VERSION : 1.0
// Support: tech.team.motioncontrol@siemens.com
   VAR_INPUT
      Cfg_EventListOffset : Int;   // Commanded event list offset (used for scrolling)
      Cfg_FilterCategory : Int;   // Filtered category number
      Cfg_TimeSortDirection : Bool;   // 1=newest first; 0=oldest first
      Cmd_FilterActiveEvents : Bool;   // 1=only show active events; 0=show all events
      Cmd_FilterCategory : Bool;   // Filter events to show only selected category number
      Cmd_SortCategory : Bool;   // 1=Sort events by ascending category number
   END_VAR
   VAR_OUTPUT
      Sts_EventListOffset : Int;   // Actual event list offset
      Sts_FilterExcludedNumEvents : Int;   // The number of events excluded by filtering
      Sts_SortFilterNumEvents : Int;   // Number of events in the sorted or filtered event list
   END_VAR
   VAR_IN_OUT
      In_Events : Array[0.."CPG_NO_OF_STS_ELEMENTS_EVENT_SUM_UPPER_LIM"] of "CPG_typeEvent";   // Input Event list to be sorted and/or filtered
      In_NumEvents : Int;   // Number of events to be sorted and/or filtered
      Sts_SortFilterEventList : Array[0.."CPG_NO_OF_HMI_SORT_EVENTS_UPPER_LIM"] of "CPG_typeEvent";   // Output sorted and/or filtered event list
   END_VAR
   VAR
      statFirstScan : Bool;   // stat first scan bit
      statCatIndex : Int;   // stat category index
      statCopiedIndex : Int;   // stat copied index
      statFilterActive : Bool;   // stat filter active = 1
      statFilterCategory : Bool;   // stat filter category
      statFilteredIndex : Int;   // stat filtered index
      statIndex : Int;   // stat index
      statLocalEventOffset : Int;   // stat local event offset
      statMaxInputSize : Int;   // stat max input size
      statMaxLocalInputSize : Int;   // stat max local input size
      statMaxOutputSize : Int;   // stat max output size
      statMaxParameterInputSize : Int;   // stat max parameter input size
      statNumDisplayedEvents : Int;   // stat num displayed events
      statNumFilteredEvents : Int;   // stat num of filtered events
      statPrevNumEvents : Int;   // stat previous number of events
      statSortedIndex : Int;   // stat sorted index
      statFilteredEventList : Array[0.."CPG_NO_OF_STS_ELEMENTS_EVENT_SUM_UPPER_LIM"] of "CPG_typeEvent";   // stat sorted event list
      statZeroEvent : "CPG_typeEvent";   // stat zeroized event list
   END_VAR
   VAR_TEMP
      tempMoveBlkVariantRetVal : Int;   // temp return value for BlockMoveVariant
   END_VAR
   VAR CONSTANT
      ZERO_VALUE : Int := 0;
   END_VAR
BEGIN
   //============================================================================================================
   // SIEMENS AG
   // (c)Copyright 2018 All Rights Reserved
   //------------------------------------------------------------------------------------------------------------
   // Project: CPG Template
   // Tested with: S7-1500 with FW version V2.1
   // Engineering: TIA Portal V14
   // Restrictions: ---
   // Requirements: S7-1500
   // Functionality: Control Event Sort Filter commands
   // Support: tech.team.motioncontrol@siemens.com
   //------------------------------------------------------------------------------------------------------------
   // Change log table:
   // Version       Date               Expert in charge    Changes applied
   //  01.00.00     01.01.2018         MP                  Initial Release & PackML V2.1  Renamed CPG V1.0
   //  01.01.00     29.05.2018         JP                  Adopted to styleguide
   //============================================================================================================
   // Function : CPG_EventSortFilter
   //============================================================================================================

   IF #statFirstScan = FALSE THEN
       // initialize & determine max array size
       // input array size (i.e. Array[0.."CPG_NO_STS_ELEMENTS_EVENT_STATUS"] of "typeCPG_Event")
       "CPG_ArrayLength"(arrayToBeSized := #In_Events,
                         arraySize => #statMaxParameterInputSize);

       //output array size for HMI (i.e. Array[0.."CPG_NO_HMI_SORT_EVENTS"] of "typeCPG_Event")
       "CPG_ArrayLength"(arrayToBeSized := #Sts_SortFilterEventList,
                         arraySize => #statMaxOutputSize);

       // internal/temporary array size (i.e. Array[0.."CPG_NO_STS_ELEMENTS_EVENT_STATUS"] of "typeCPG_Event")   
       "CPG_ArrayLength"(arrayToBeSized := #statFilteredEventList,
                                 arraySize => #statMaxLocalInputSize);

       //Take smallest aray as the maximum number of input events to filter and sort
       IF #statMaxParameterInputSize > #statMaxLocalInputSize THEN
           #statMaxInputSize := #statMaxLocalInputSize;
       ELSE
           #statMaxInputSize := #statMaxParameterInputSize;
       END_IF;
       // clear the output sort buffer
       FOR #statIndex := 0 TO #statMaxOutputSize - 1 DO
           #Sts_SortFilterEventList[#statIndex] := #statZeroEvent;
       END_FOR;

       #statFirstScan := TRUE;            // set the first scan bit 
   END_IF;
   // End of First Scan Section


   // Main Filter Logic

   #statFilteredIndex := 0;
   // sort by ascending OR descending?
   IF #Cfg_TimeSortDirection THEN
       #statIndex := #In_NumEvents - 1;  // newest events first
   ELSE
       #statIndex := 0;   // oldest events first
   END_IF;

   IF #In_NumEvents > 0 THEN

       REPEAT
           #statFilterCategory := 0;
           #statFilterActive := 0;
           IF #Cmd_FilterCategory AND (#In_Events[#statIndex].Category = #Cfg_FilterCategory) THEN
               #statFilterCategory := 1;
           END_IF;
           IF #Cmd_FilterActiveEvents AND (#In_Events[#statIndex].Trigger) THEN
               #statFilterActive := 1;
           END_IF;

           IF ((#Cmd_FilterCategory AND #statFilterCategory) OR NOT (#Cmd_FilterCategory)) AND ((#Cmd_FilterActiveEvents AND #statFilterActive) OR NOT (#Cmd_FilterActiveEvents)) THEN
               #statFilteredEventList[#statFilteredIndex] := #In_Events[#statIndex];
               #statFilteredIndex := #statFilteredIndex + 1;
           END_IF;

           IF #Cfg_TimeSortDirection THEN
               #statIndex := #statIndex - 1;
           ELSE
               #statIndex := #statIndex + 1;
           END_IF;

       UNTIL #statFilteredIndex >= #In_NumEvents OR #statFilteredIndex >= #statMaxInputSize OR #statIndex < 0 OR #statIndex >= #In_NumEvents END_REPEAT;
   END_IF;

   #statNumFilteredEvents := #statFilteredIndex;

   #Sts_SortFilterNumEvents := #statNumFilteredEvents;
   #Sts_FilterExcludedNumEvents := #In_NumEvents - #statNumFilteredEvents;

   //Sanitize and limit Cfg_EventListOffset, offset cannot go past the last event
   IF #Cfg_EventListOffset > #statNumFilteredEvents - 1 THEN
       #statLocalEventOffset := #statNumFilteredEvents - 1;
   ELSE
       #statLocalEventOffset := #Cfg_EventListOffset;
   END_IF;

   IF #statLocalEventOffset < 0 THEN
       #statLocalEventOffset := 0;
   END_IF;
   #Sts_EventListOffset := #statLocalEventOffset;

   #statSortedIndex := 0;
   #statCopiedIndex := 0;

   //Category sorting loops
   IF #Cmd_SortCategory THEN
       IF #statNumFilteredEvents <> 0 THEN
           #statCatIndex := 0;
           REPEAT //Repeat for categories 0-9
               #statIndex := 0;

               REPEAT //Repeat for every event in the filtered list
                   //If the category matches, add to the list

                   IF #statCatIndex = #statFilteredEventList[#statIndex].Category THEN
                       //Track sorted index separate from copied index.  
                       //This allows a "hypothetical" sort when an offset is applied, without using memory for a non-offset sorted list
                       IF (#statSortedIndex >= #statLocalEventOffset) THEN
                           #Sts_SortFilterEventList[#statCopiedIndex] := #statFilteredEventList[#statIndex];
                           #statCopiedIndex := #statCopiedIndex + 1;
                       END_IF;
                       #statSortedIndex := #statSortedIndex + 1;
                   END_IF;

                   IF #statCopiedIndex >= #statMaxOutputSize THEN
                       EXIT; //EXIT unsorted loop
                   END_IF;

                   #statIndex := #statIndex + 1;
               UNTIL #statIndex >= #statNumFilteredEvents END_REPEAT;

               IF #statCopiedIndex >= #statMaxOutputSize THEN
                   EXIT; //EXIT category loop
               END_IF;
               #statCatIndex := #statCatIndex + 1;
           UNTIL #statCatIndex > 9 END_REPEAT;

           //Handle display of events in the case the category is not 0-9, but do not sort in order for scan time purposes
           //Only for special cases
           IF #statCopiedIndex < #statMaxOutputSize - 1 AND #statSortedIndex <> #statNumFilteredEvents THEN
               #statIndex := 0;
               REPEAT
                   IF #statFilteredEventList[#statIndex].Category > 9 THEN
                       IF (#statSortedIndex >= #statLocalEventOffset) THEN
                           #Sts_SortFilterEventList[#statCopiedIndex] := #statFilteredEventList[#statIndex];
                           #statCopiedIndex := #statCopiedIndex + 1;
                       END_IF;

                       #statSortedIndex := #statSortedIndex + 1;

                   END_IF;


                   IF #statCopiedIndex >= #statMaxOutputSize THEN
                       EXIT;
                   END_IF;

                   #statIndex := #statIndex + 1;

               UNTIL #statIndex >= #statNumFilteredEvents END_REPEAT;

           END_IF;

       END_IF;

   ELSE
       //If no category sorting is done, copy the entire filtered list and apply any offset
       #statCopiedIndex := #statNumFilteredEvents - #statLocalEventOffset;

       IF #statCopiedIndex > #statMaxOutputSize THEN
           #statCopiedIndex := #statMaxOutputSize;
       ELSIF #statCopiedIndex < 0 THEN
           #statCopiedIndex := 0;
       END_IF;

       #tempMoveBlkVariantRetVal := MOVE_BLK_VARIANT(SRC := #statFilteredEventList, COUNT := DINT_TO_UDINT(#statCopiedIndex), SRC_INDEX := #statLocalEventOffset, DEST_INDEX := #ZERO_VALUE, DEST => #Sts_SortFilterEventList);

   END_IF;

   #statNumDisplayedEvents := #statCopiedIndex;

   // Clean up event list
   IF #statPrevNumEvents > #statNumDisplayedEvents THEN
       FOR #statIndex := #statNumDisplayedEvents TO #statPrevNumEvents - 1 DO
           #Sts_SortFilterEventList[#statIndex] := #statZeroEvent;
       END_FOR;
   END_IF;

   #statPrevNumEvents := #statNumDisplayedEvents;

   //  -------------- END OF LOGIC -------------------------
   ENO := TRUE;   // Set the ENO output
END_FUNCTION_BLOCK

FUNCTION_BLOCK "CPG_EventSummation"   // FB31605, SCL
TITLE = CPG_EventSummation
{ S7_Optimized_Access := 'TRUE' }
AUTHOR : tech.team.motioncontrol@siemens.com
FAMILY : CPG
VERSION : 1.0
// Support: tech.team.motioncontrol@siemens.com
   VAR_OUTPUT
      Sts_NumEvents : Int;   // Status - Number of active events
      Sts_Category_0_Latched : Bool;   // Status - Latched Event - Cat. 0
      Sts_Category_1_Latched : Bool;   // Status - Latched Event - Cat. 1
      Sts_Category_2_Latched : Bool;   // Status - Latched Event - Cat. 2
      Sts_Category_3_Latched : Bool;   // Status - Latched Event - Cat. 3
      Sts_Category_4_Latched : Bool;   // Status - Latched Event - Cat. 4
      Sts_Category_5_Latched : Bool;   // Status - Latched Event - Cat. 5
      Sts_Category_6_Latched : Bool;   // Status - Latched Event - Cat. 6
      Sts_Category_7_Latched : Bool;   // Status - Latched Event - Cat. 7
      Sts_Category_8_Latched : Bool;   // Status - Latched Event - Cat. 8
      Sts_Category_9_Latched : Bool;   // Status - Latched Event - Cat. 9
      Sts_Category_0_NotLatched : Bool;   // Status - NotLatched (Active) Event - Cat. 0
      Sts_Category_1_NotLatched : Bool;   // Status - NotLatched (Active) Event - Cat. 1
      Sts_Category_2_NotLatched : Bool;   // Status - NotLatched (Active) Event - Cat. 2
      Sts_Category_3_NotLatched : Bool;   // Status - NotLatched (Active) Event - Cat. 3
      Sts_Category_4_NotLatched : Bool;   // Status - NotLatched (Active) Event - Cat. 4
      Sts_Category_5_NotLatched : Bool;   // Status - NotLatched (Active) Event - Cat. 5
      Sts_Category_6_NotLatched : Bool;   // Status - NotLatched (Active) Event - Cat. 6
      Sts_Category_7_NotLatched : Bool;   // Status - NotLatched (Active) Event - Cat. 7
      Sts_Category_8_NotLatched : Bool;   // Status - NotLatched (Active) Event - Cat. 8
      Sts_Category_9_NotLatched : Bool;   // Status - NotLatched (Active) Event - Cat. 9
      Sts_CurrentActiveEvent : Bool;   // Active Event Exists
      Sts_Error : Bool;   // Error in FB
      Sts_ErrorCode : DInt;   // Error Code
   END_VAR
   VAR_IN_OUT
      In_EventStatus : "CPG_typeEventStatus";   // UDT of EventStatus
      Sts_EventSummation : "CPG_typeEventSummation";   // UDT of EventSummation
   END_VAR
   VAR
      statFirstScan : Bool;   // 0=1st scan of FB; set to 1 after 1st FB scan...
      statCfg_MaxEvents : Int;   // number of events used from In_EventStatus array.
      statEventsRemaining : Int;   // number of events remaining
      statCompareTrue : Bool;   // Compare true?
      statIndex : Int;   // Index counter
      statIndex1 : Int;   // Index counter
      statIndex2 : Int;   // Index counter
      statIndex3 : Int;   // Index counter
      statIndex3a : Int;   // Index counter
      statIndex3AOffset : Int;   // Index counter
      statWriteData : Bool;
   END_VAR
   VAR_TEMP
      tempDTL1 : DTL;   // Temp Date & Time value as DTL format
      tempDTL2 : DTL;   // Temp Date & Time value as DTL format
      tempMoveBlkVariantRetVal : Int;   // temp return value for BlockMoveVariant
   END_VAR
BEGIN
   //============================================================================================================
   // SIEMENS AG
   // (c)Copyright 2018 All Rights Reserved
   //------------------------------------------------------------------------------------------------------------
   // Project: CPG Template
   // Tested with: S7-1500 with FW version V2.1
   // Engineering: TIA Portal V14
   // Restrictions: ---
   // Requirements: S7-1500
   // Functionality:  Summarizes the "Data" from the equipment modules (from FB_EventManager) AND will create one list OF events FOR the unit machine.
   //                 It summarizes the data by finding the unit machine first out event and summarizes which category of events are active.
   //                 CPG_EventSummationBegin initializes the summation, and CPG_EventSummationEnd finalizes the summation.
   // Support: tech.team.motioncontrol@siemens.com
   //------------------------------------------------------------------------------------------------------------
   // Change log table:
   // Version       Date               Expert in charge    Changes applied
   //  01.00.00     01.01.2018         MP                  Initial Release & PackML V2.1  Renamed CPG V1.0
   //  01.01.00     29.05.2018         JP                  Adopted to styleguide
   //============================================================================================================
   // Function Block : CPG_EventSummation
   //============================================================================================================


   // ===========================================================================
   //  BEGIN THE LOGIC SECTION:
   //  First scan section
   IF #statFirstScan = FALSE THEN
       // initialize & determine max array size
       // input array size (i.e. Array[0.."CPG_NO_STS_ELEMENTS_EVENT_STATUS"] of "typeCPG_Event")
       "CPG_ArrayLength"(arrayToBeSized := #In_EventStatus.sts_Events,
                         arraySize => #In_EventStatus.wrk_EventArraySize);

       "CPG_ArrayLength"(arrayToBeSized := #In_EventStatus.sts_Events,
                         arraySize => #statCfg_MaxEvents);

       #statFirstScan := TRUE;            // set the first scan bit 
   END_IF;
   // End of First Scan Section


   // BEGIN THE MAIN LOGIC SECTION:
   #Sts_ErrorCode := 0;               // Set the status error code
   #statWriteData := FALSE;                // set write data to false

   // Set First Out Event
   #tempDTL1 := #In_EventStatus.sts_FirstOutEvent.DateTimeDTL;                  // Date & Time of Sts_FirstOutEventCat[index].TimeEvent

   IF #tempDTL1 <> DTL#1970-01-01-00:00:00.0 THEN                                  // is In_EventStatus.Sts_FirstOutEvent.TimeEvent <> 0?
      #tempDTL2 := #Sts_EventSummation.sts_FirstOutEvent.DateTimeDTL;           // load the current value of the Sts_Eve..
      #statWriteData := FALSE;                                                   // Reset the write data command.
         IF #tempDTL2 = DTL#1970-01-01-00:00:00.0 THEN                             // is Sts_EventSummation.Sts_FirstOutEvent.TimeEvent = 0? 
              #statWriteData := TRUE;
         ELSIF #tempDTL1 < #tempDTL2 THEN                                   // is IN_event newer than Sts_event ?
             #statWriteData := TRUE;
         END_IF;     // End "IF (EQ_DT(DT1:=Sts_"
   END_IF;         // End "IF (NOT(EQ_DT(DT1:=In_Ev"

   IF #statWriteData THEN 
      #Sts_EventSummation.sts_FirstOutEvent := #In_EventStatus.sts_FirstOutEvent;  // Update the First Fault event 
   END_IF; 

   // Set First Out Event by Category
   FOR #statIndex:= 0 TO 9 DO

       #tempDTL1:=#In_EventStatus.sts_FirstOutEventCat[#statIndex].DateTimeDTL;        // Date & Time of Sts_FirstOutEventCat[index].TimeEvent

       IF #tempDTL1 <> DTL#1970-01-01-00:00:00.0 THEN                                // is In_EventStatus.Sts_FirstOutEvent.TimeEvent <> 0?

           #tempDTL2:=#Sts_EventSummation.sts_FirstOutEventCat[#statIndex].DateTimeDTL;          // load the current value of the Sts_Eve..
           #statWriteData:=0;                   // Reset the write data command.

           IF #tempDTL2 = DTL#1970-01-01-00:00:00.0 THEN                              // is Sts_EventSummation.Sts_FirstOutEvent.TimeEvent = 0? 
               #statWriteData := TRUE;

           ELSIF #tempDTL1 < #tempDTL2 THEN   // is IN_event newer than Sts_event ?

               #statWriteData := TRUE;

           END_IF;     // End "IF (EQ_DT(DT1:=Sts_"
       END_IF;         // End "IF (NOT(EQ_DT(DT1:=In_Ev"

       IF #statWriteData THEN 
           #Sts_EventSummation.sts_FirstOutEventCat[#statIndex] := #In_EventStatus.sts_FirstOutEventCat[#statIndex];  // Update the First Fault event 
       END_IF; 
   END_FOR;     

   // ---------------------------------------------------------------
   // Set Active Events
   IF #In_EventStatus.sts_NumEvents > 0 THEN 
       IF #In_EventStatus.sts_NumEvents > 0 AND #Sts_EventSummation.sts_NumEvents > 0 THEN
           #statIndex1 := 0;
           FOR #statIndex := 0 TO #In_EventStatus.sts_NumEvents - 1 DO

               WHILE #statIndex1 < #Sts_EventSummation.sts_NumEvents DO

                   #statCompareTrue := FALSE;
                   #statIndex2 := 0;

                   REPEAT
                       IF #In_EventStatus.sts_Events[#statIndex].DateTimeDTL = #Sts_EventSummation.sts_Events[#statIndex1].DateTimeDTL THEN
                           #statIndex2 := #statIndex2 + 1;

                       ELSIF #In_EventStatus.sts_Events[#statIndex].DateTimeDTL < #Sts_EventSummation.sts_Events[#statIndex1].DateTimeDTL THEN
                           #statCompareTrue := TRUE;

                           EXIT;  // Exit the REPEAT loop
                       ELSE
                           EXIT;  // Exit the REPEAT loop
                       END_IF;
                   UNTIL #statIndex2 = 7
                   END_REPEAT;

                   IF #statCompareTrue THEN
                       #statEventsRemaining := #Sts_EventSummation.sts_NumEvents - #statIndex1;
                       #statIndex3AOffset := #statEventsRemaining - 1 + #statIndex1;

                       FOR #statIndex3 := 0 TO #statEventsRemaining - 1 DO  // Backwards copy the data to shift it down to prevent the data from overwriting itself
                           #statIndex3a := #statIndex3AOffset - #statIndex3;
                           IF #statIndex3a + 1 < #Sts_EventSummation.wrk_EventArraySize THEN
                               #Sts_EventSummation.sts_Events[#statIndex3a + 1] := #Sts_EventSummation.sts_Events[#statIndex3a];
                           END_IF;
                       END_FOR;

                       #Sts_EventSummation.sts_Events[#statIndex1] := #In_EventStatus.sts_Events[#statIndex];

                       IF #Sts_EventSummation.sts_NumEvents < #Sts_EventSummation.wrk_EventArraySize THEN
                           #Sts_EventSummation.sts_NumEvents := #Sts_EventSummation.sts_NumEvents + 1;
                           #statIndex1 := #statIndex1 + 1;
                       END_IF;

                       EXIT;  //Exit the WHILE loop
                   END_IF;
                   #statIndex1 := #statIndex1 + 1;
               END_WHILE;

               // If the WHILE loop is done, then bulk copy the remaining events into the event summation array.
               IF #statIndex1 = #Sts_EventSummation.sts_NumEvents THEN
                   #statEventsRemaining := #In_EventStatus.sts_NumEvents - #statIndex;
                   IF #statEventsRemaining + #Sts_EventSummation.sts_NumEvents > #Sts_EventSummation.wrk_EventArraySize THEN
                       #statEventsRemaining := #Sts_EventSummation.wrk_EventArraySize - #Sts_EventSummation.sts_NumEvents;
                       #Sts_ErrorCode := 1;
                   END_IF;

                   IF #statEventsRemaining > 0 THEN
                       #Sts_EventSummation.sts_Events[#statIndex1] := #In_EventStatus.sts_Events[#statIndex];
                       #Sts_EventSummation.sts_NumEvents := #Sts_EventSummation.sts_NumEvents + #statEventsRemaining;
                   END_IF;
                   EXIT;  //Exit the FOR loop
               END_IF;
           END_FOR;
       ELSIF #In_EventStatus.sts_NumEvents > 0 THEN
           // The current event summation array is empty, so just bulk copy the data over.
           IF #In_EventStatus.sts_NumEvents < #Sts_EventSummation.wrk_EventArraySize THEN

               #tempMoveBlkVariantRetVal := MOVE_BLK_VARIANT(SRC := #In_EventStatus.sts_Events,
                                                                    COUNT := INT_TO_UDINT(#In_EventStatus.sts_NumEvents),
                                                                    SRC_INDEX := 0,
                                                                    DEST_INDEX := 0,
                                                                    DEST => #Sts_EventSummation.sts_Events);
               #Sts_EventSummation.sts_NumEvents := #In_EventStatus.sts_NumEvents;
           ELSE

               #tempMoveBlkVariantRetVal := MOVE_BLK_VARIANT(SRC := #In_EventStatus.sts_Events,
                                                                    COUNT := INT_TO_UDINT (#Sts_EventSummation.wrk_EventArraySize),
                                                                    SRC_INDEX := 0,
                                                                    DEST_INDEX := 0,
                                                                    DEST => #Sts_EventSummation.sts_Events);
               #Sts_EventSummation.sts_NumEvents := #Sts_EventSummation.wrk_EventArraySize;
               #Sts_ErrorCode := 1;
           END_IF;


       END_IF;    
   END_IF;

   // update the output
   #Sts_NumEvents := #Sts_EventSummation.sts_NumEvents;

   // Set Category Bits
   #Sts_EventSummation.wrk_Category_0_Latched := (#Sts_EventSummation.wrk_Category_0_Latched OR #In_EventStatus.sts_Category_0_Latched);
   #Sts_EventSummation.wrk_Category_1_Latched := (#Sts_EventSummation.wrk_Category_1_Latched OR #In_EventStatus.sts_Category_1_Latched);
   #Sts_EventSummation.wrk_Category_2_Latched := (#Sts_EventSummation.wrk_Category_2_Latched OR #In_EventStatus.sts_Category_2_Latched);
   #Sts_EventSummation.wrk_Category_3_Latched := (#Sts_EventSummation.wrk_Category_3_Latched OR #In_EventStatus.sts_Category_3_Latched);
   #Sts_EventSummation.wrk_Category_4_Latched := (#Sts_EventSummation.wrk_Category_4_Latched OR #In_EventStatus.sts_Category_4_Latched);
   #Sts_EventSummation.wrk_Category_5_Latched := (#Sts_EventSummation.wrk_Category_5_Latched OR #In_EventStatus.sts_Category_5_Latched);
   #Sts_EventSummation.wrk_Category_6_Latched := (#Sts_EventSummation.wrk_Category_6_Latched OR #In_EventStatus.sts_Category_6_Latched);
   #Sts_EventSummation.wrk_Category_7_Latched := (#Sts_EventSummation.wrk_Category_7_Latched OR #In_EventStatus.sts_Category_7_Latched);
   #Sts_EventSummation.wrk_Category_8_Latched := (#Sts_EventSummation.wrk_Category_8_Latched OR #In_EventStatus.sts_Category_8_Latched);
   #Sts_EventSummation.wrk_Category_9_Latched := (#Sts_EventSummation.wrk_Category_9_Latched OR #In_EventStatus.sts_Category_9_Latched);

   #Sts_Category_0_Latched := #In_EventStatus.sts_Category_0_Latched;
   #Sts_Category_1_Latched := #In_EventStatus.sts_Category_1_Latched;
   #Sts_Category_2_Latched := #In_EventStatus.sts_Category_2_Latched;
   #Sts_Category_3_Latched := #In_EventStatus.sts_Category_3_Latched;
   #Sts_Category_4_Latched := #In_EventStatus.sts_Category_4_Latched;
   #Sts_Category_5_Latched := #In_EventStatus.sts_Category_5_Latched;
   #Sts_Category_6_Latched := #In_EventStatus.sts_Category_6_Latched;
   #Sts_Category_7_Latched := #In_EventStatus.sts_Category_7_Latched;
   #Sts_Category_8_Latched := #In_EventStatus.sts_Category_8_Latched;
   #Sts_Category_9_Latched := #In_EventStatus.sts_Category_9_Latched;

   #Sts_EventSummation.wrk_Category_0_NotLatched := #Sts_EventSummation.wrk_Category_0_NotLatched OR #In_EventStatus.sts_Category_0_NotLatched;
   #Sts_EventSummation.wrk_Category_1_NotLatched := #Sts_EventSummation.wrk_Category_1_NotLatched OR #In_EventStatus.sts_Category_1_NotLatched;
   #Sts_EventSummation.wrk_Category_2_NotLatched := #Sts_EventSummation.wrk_Category_2_NotLatched OR #In_EventStatus.sts_Category_2_NotLatched;
   #Sts_EventSummation.wrk_Category_3_NotLatched := #Sts_EventSummation.wrk_Category_3_NotLatched OR #In_EventStatus.sts_Category_3_NotLatched;
   #Sts_EventSummation.wrk_Category_4_NotLatched := #Sts_EventSummation.wrk_Category_4_NotLatched OR #In_EventStatus.sts_Category_4_NotLatched;
   #Sts_EventSummation.wrk_Category_5_NotLatched := #Sts_EventSummation.wrk_Category_5_NotLatched OR #In_EventStatus.sts_Category_5_NotLatched;
   #Sts_EventSummation.wrk_Category_6_NotLatched := #Sts_EventSummation.wrk_Category_6_NotLatched OR #In_EventStatus.sts_Category_6_NotLatched;
   #Sts_EventSummation.wrk_Category_7_NotLatched := #Sts_EventSummation.wrk_Category_7_NotLatched OR #In_EventStatus.sts_Category_7_NotLatched;
   #Sts_EventSummation.wrk_Category_8_NotLatched := #Sts_EventSummation.wrk_Category_8_NotLatched OR #In_EventStatus.sts_Category_8_NotLatched;
   #Sts_EventSummation.wrk_Category_9_NotLatched := #Sts_EventSummation.wrk_Category_9_NotLatched OR #In_EventStatus.sts_Category_9_NotLatched;

   #Sts_Category_0_NotLatched := #In_EventStatus.sts_Category_0_NotLatched;
   #Sts_Category_1_NotLatched := #In_EventStatus.sts_Category_1_NotLatched;
   #Sts_Category_2_NotLatched := #In_EventStatus.sts_Category_2_NotLatched;
   #Sts_Category_3_NotLatched := #In_EventStatus.sts_Category_3_NotLatched;
   #Sts_Category_4_NotLatched := #In_EventStatus.sts_Category_4_NotLatched;
   #Sts_Category_5_NotLatched := #In_EventStatus.sts_Category_5_NotLatched;
   #Sts_Category_6_NotLatched := #In_EventStatus.sts_Category_6_NotLatched;
   #Sts_Category_7_NotLatched := #In_EventStatus.sts_Category_7_NotLatched;
   #Sts_Category_8_NotLatched := #In_EventStatus.sts_Category_8_NotLatched;
   #Sts_Category_9_NotLatched := #In_EventStatus.sts_Category_9_NotLatched;

   #Sts_EventSummation.wrk_CurrentActiveEvent := #Sts_EventSummation.wrk_CurrentActiveEvent OR #In_EventStatus.sts_CurrentActiveEvent;

   #Sts_CurrentActiveEvent := #In_EventStatus.sts_CurrentActiveEvent;

   // Set Error Bit
   #Sts_Error := (#Sts_ErrorCode <> 0);

   //  -------------- END OF LOGIC -------------------------
   ENO := TRUE;   // Set the ENO output
END_FUNCTION_BLOCK

FUNCTION_BLOCK "CPG_EventSummationBegin"   // FB31606, SCL
TITLE = CPG_EventSummationBegin
{ S7_Optimized_Access := 'TRUE' }
AUTHOR : tech.team.motioncontrol@siemens.com
FAMILY : CPG
VERSION : 1.0
// Support: tech.team.motioncontrol@siemens.com
   VAR_IN_OUT
      Sts_EventSummation : "CPG_typeEventSummation";   // Working event list data section
   END_VAR
   VAR
      statFirstScan : Bool;   // 0=1st scan of FB; set to 1 after 1st FB scan...
      statIndex : Int;   // temp value needed with FOR loop
      statZeroEvent : "CPG_typeEvent";   // Null Event
   END_VAR
BEGIN
   //============================================================================================================
   // SIEMENS AG
   // (c)Copyright 2018 All Rights Reserved
   //------------------------------------------------------------------------------------------------------------
   // Project: CPG Template
   // Tested with: S7-1500 with FW version V2.1
   // Engineering: TIA Portal V14
   // Restrictions: ---
   // Requirements: S7-1500
   // Functionality:  Summarizes the "Data" from the equipment modules (from FB_EventManager) AND will create one list OF events FOR the unit machine.
   //                 It summarizes the data by finding the unit machine first out event and summarizes which category of events are active.
   //                 FB_EventSummationBegin initializes the summation, and FB_EventSummationEnd finalizes the summation.
   // Support: tech.team.motioncontrol@siemens.com
   //------------------------------------------------------------------------------------------------------------
   // Change log table:
   // Version       Date               Expert in charge    Changes applied
   //  01.00.00     01.01.2018         MP                  Initial Release & PackML V2.1  Renamed CPG V1.0
   //  01.01.00     29.05.2018         JP                  Adopted to styleguide
   //============================================================================================================
   // Function Block : CPG_EventSummationBegin
   //============================================================================================================



   // ===========================================================================
   // Begin the First Scan / Initialize logic section:
   IF #statFirstScan = FALSE THEN
       // initialize & determine max array size
       "CPG_ArrayLength"(arrayToBeSized := #Sts_EventSummation.sts_Events,
                         arraySize => #Sts_EventSummation.wrk_EventArraySize);

       // initialize and clear the status events area
              FOR #statIndex := 0 TO (#Sts_EventSummation.wrk_EventArraySize - 1) DO
                  #Sts_EventSummation.sts_Events[#statIndex] := #statZeroEvent;
              END_FOR;

       #statFirstScan := TRUE;            // set the first scan bit 
   END_IF;
   // End of First Scan Section

   // Begin the LOGIC section:
   // Initialize the summation - This FB is to be called before the numerous "FB_PG_EventSum" calls.

   // Clear the first out event
   #Sts_EventSummation.sts_FirstOutEvent := #statZeroEvent;

   // Clear the first out event category arrays  
   FOR #statIndex := 0 TO 9 DO
       #Sts_EventSummation.sts_FirstOutEventCat[#statIndex] := #statZeroEvent;
   END_FOR;

   // Determine the array size
   "CPG_ArrayLength"(arrayToBeSized := #Sts_EventSummation.sts_Events,
                            arraySize => #Sts_EventSummation.wrk_EventArraySize);
   // Clear the number of events
   #Sts_EventSummation.sts_NumEvents := 0;            // set the number of events to 0.

   // Clear the output category status bits
   #Sts_EventSummation.wrk_Category_0_Latched := FALSE;
   #Sts_EventSummation.wrk_Category_1_Latched := FALSE;
   #Sts_EventSummation.wrk_Category_2_Latched := FALSE;
   #Sts_EventSummation.wrk_Category_3_Latched := FALSE;
   #Sts_EventSummation.wrk_Category_4_Latched := FALSE;
   #Sts_EventSummation.wrk_Category_5_Latched := FALSE;
   #Sts_EventSummation.wrk_Category_6_Latched := FALSE;
   #Sts_EventSummation.wrk_Category_7_Latched := FALSE;
   #Sts_EventSummation.wrk_Category_8_Latched := FALSE;
   #Sts_EventSummation.wrk_Category_9_Latched := FALSE;
   #Sts_EventSummation.wrk_Category_0_NotLatched := FALSE;
   #Sts_EventSummation.wrk_Category_1_NotLatched := FALSE;
   #Sts_EventSummation.wrk_Category_2_NotLatched := FALSE;
   #Sts_EventSummation.wrk_Category_3_NotLatched := FALSE;
   #Sts_EventSummation.wrk_Category_4_NotLatched := FALSE;
   #Sts_EventSummation.wrk_Category_5_NotLatched := FALSE;
   #Sts_EventSummation.wrk_Category_6_NotLatched := FALSE;
   #Sts_EventSummation.wrk_Category_7_NotLatched := FALSE;
   #Sts_EventSummation.wrk_Category_8_NotLatched := FALSE;
   #Sts_EventSummation.wrk_Category_9_NotLatched := FALSE;
   #Sts_EventSummation.wrk_CurrentActiveEvent := FALSE;

   //  -------------- END OF LOGIC -------------------------
   ENO := TRUE;   // Set the ENO output
END_FUNCTION_BLOCK

FUNCTION_BLOCK "CPG_EventSummationEnd"   // FB31607, SCL
TITLE = CPG_EventSummationEnd
{ S7_Optimized_Access := 'TRUE' }
AUTHOR : tech.team.motioncontrol@siemens.com
FAMILY : CPG
VERSION : 1.0
// Support: tech.team.motioncontrol@siemens.com
   VAR_IN_OUT
      Sts_EventSummation : "CPG_typeEventSummation";   // Working event list data section
   END_VAR
   VAR
      statFirstScan : Bool;   // 0=1st scan of FB; set to 1 after 1st FB scan...
      statIndex : Int;   // stat index
      statPrev_NumAllEvents : Int;   // stat value needed with FOR loop
   END_VAR
   VAR_TEMP
      tempZeroEvent : "CPG_typeEvent";   // null instance of UDT Event
   END_VAR
BEGIN
   //============================================================================================================
   // SIEMENS AG
   // (c)Copyright 2018 All Rights Reserved
   //------------------------------------------------------------------------------------------------------------
   // Project: CPG Template
   // Tested with: S7-1500 with FW version V2.1
   // Engineering: TIA Portal V14
   // Restrictions: ---
   // Requirements: S7-1500
   // Functionality:  Summarizes the "Data" from the equipment modules (from FB_EventManager) AND will create one list OF events FOR the unit machine.
   //                 It summarizes the data by finding the unit machine first out event and summarizes which category of events are active.
   //                 CPG_EventSummationBegin initializes the summation, and CPG_EventSummationEnd finalizes the summation.
   // Support: tech.team.motioncontrol@siemens.com
   //------------------------------------------------------------------------------------------------------------
   // Change log table:
   // Version       Date               Expert in charge    Changes applied
   //  01.00.00     01.01.2018         MP                  Initial Release & PackML V2.1  Renamed CPG V1.0
   //  01.01.00     29.05.2018         JP                  Adopted to styleguide
   //  01.00.01     13.06.2019         ThH                 Corrected handling of Bit 5; new Version CPG Template V1.0.1
   //============================================================================================================
   // Function Block : CPG_EventSummationEnd
   //============================================================================================================

   // ===========================================================================
   //  Begin the LOGIC section:
   // first scan logic
   IF #statFirstScan = FALSE THEN
       // initialize & determine max array size
       "CPG_ArrayLength"(arrayToBeSized := #Sts_EventSummation.sts_Events,
                         arraySize => #Sts_EventSummation.wrk_EventArraySize);

       #statPrev_NumAllEvents := #Sts_EventSummation.wrk_EventArraySize;

       #statFirstScan := TRUE;            // set the first scan bit
   END_IF;

   // Cleanup the summation - This FB is to be called after the numerous "FB_PMLe_EventSum" calls.
   IF #statPrev_NumAllEvents > #Sts_EventSummation.sts_NumEvents THEN

       FOR #statIndex := #Sts_EventSummation.sts_NumEvents TO (#statPrev_NumAllEvents-1) DO
           #Sts_EventSummation.sts_Events[#statIndex]:= #tempZeroEvent;   // clear event area of cleared alarms
       END_FOR;

   END_IF;

   #statPrev_NumAllEvents := #Sts_EventSummation.sts_NumEvents;     

   // Update the output bits from work area
   #Sts_EventSummation.sts_Category_0_Latched := #Sts_EventSummation.wrk_Category_0_Latched;
   #Sts_EventSummation.sts_Category_1_Latched := #Sts_EventSummation.wrk_Category_1_Latched;
   #Sts_EventSummation.sts_Category_2_Latched := #Sts_EventSummation.wrk_Category_2_Latched;
   #Sts_EventSummation.sts_Category_3_Latched := #Sts_EventSummation.wrk_Category_3_Latched;
   #Sts_EventSummation.sts_Category_4_Latched := #Sts_EventSummation.wrk_Category_4_Latched;
   #Sts_EventSummation.sts_Category_5_Latched := #Sts_EventSummation.wrk_Category_5_Latched;
   #Sts_EventSummation.sts_Category_6_Latched := #Sts_EventSummation.wrk_Category_6_Latched;
   #Sts_EventSummation.sts_Category_7_Latched := #Sts_EventSummation.wrk_Category_7_Latched;
   #Sts_EventSummation.sts_Category_8_Latched := #Sts_EventSummation.wrk_Category_8_Latched;
   #Sts_EventSummation.sts_Category_9_Latched := #Sts_EventSummation.wrk_Category_9_Latched;

   #Sts_EventSummation.sts_Category_0_NotLatched := #Sts_EventSummation.wrk_Category_0_NotLatched;
   #Sts_EventSummation.sts_Category_1_NotLatched := #Sts_EventSummation.wrk_Category_1_NotLatched;
   #Sts_EventSummation.sts_Category_2_NotLatched := #Sts_EventSummation.wrk_Category_2_NotLatched;
   #Sts_EventSummation.sts_Category_3_NotLatched := #Sts_EventSummation.wrk_Category_3_NotLatched;
   #Sts_EventSummation.sts_Category_4_NotLatched := #Sts_EventSummation.wrk_Category_4_NotLatched;
   #Sts_EventSummation.sts_Category_5_NotLatched := #Sts_EventSummation.wrk_Category_5_NotLatched;
   #Sts_EventSummation.sts_Category_6_NotLatched := #Sts_EventSummation.wrk_Category_6_NotLatched;
   #Sts_EventSummation.sts_Category_7_NotLatched := #Sts_EventSummation.wrk_Category_7_NotLatched;
   #Sts_EventSummation.sts_Category_8_NotLatched := #Sts_EventSummation.wrk_Category_8_NotLatched;
   #Sts_EventSummation.sts_Category_9_NotLatched := #Sts_EventSummation.wrk_Category_9_NotLatched;

   #Sts_EventSummation.sts_CurrentActiveEvent  := #Sts_EventSummation.wrk_CurrentActiveEvent; 

   //  -------------- END OF LOGIC -------------------------
   ENO := TRUE;   // Set the ENO output
END_FUNCTION_BLOCK

FUNCTION_BLOCK "CPG_MsgScroll"   // FB31608, SCL
TITLE = CPG_Msg_Scroll
{ S7_Optimized_Access := 'TRUE' }
AUTHOR : tech.team.motioncontrol@siemens.com
FAMILY : CPG
VERSION : 1.0
// Support: tech.team.motioncontrol@siemens.com
   VAR_INPUT
      Trigger : Bool;   // input trigger to enable scroll logic
      NumEvents : Int;   // input value with number of active events
      In_Events : Array[0.."CPG_NO_OF_HMI_SORT_EVENTS_UPPER_LIM"] of "CPG_typeEvent";   // incoming events list
   END_VAR
   VAR_OUTPUT
      Msg_Scroll : String[40];   // message output value
   END_VAR
   VAR
      statScrollIndex : Int;   // index value for scroll logic
      statTriggerOS : Bool;   // one shot trigger
      statMaxSize : Int;   // max size
   END_VAR
   VAR_TEMP
      tempScroll_Index_Max : Int;   // max value for scroll index
   END_VAR
BEGIN
   //============================================================================================================
   // SIEMENS AG
   // (c)Copyright 2018 All Rights Reserved
   //------------------------------------------------------------------------------------------------------------
   // Project: CPG Template
   // Tested with: S7-1500 with FW version V2.1
   // Engineering: TIA Portal V14
   // Restrictions: ---
   // Requirements: S7-1500
   // Functionality:  Used to scoll messages from an array of the active events to a single string for display on the HMI
   // Support: tech.team.motioncontrol@siemens.com
   //------------------------------------------------------------------------------------------------------------
   // Change log table:
   // Version       Date               Expert in charge    Changes applied
   //  01.00.00     01.01.2018         MP                  Initial Release & PackML V2.1  Renamed CPG V1.0
   //  01.01.00     29.05.2018         JP                  Adopted to styleguide
   //============================================================================================================
   // Function Block : CPG_Msg_Scroll
   //============================================================================================================



   // ===========================================================================
   //  Begin the LOGIC section:
   // initialize & determine max array size
   "CPG_ArrayLength"(arrayToBeSized := #In_Events,
                            arraySize => #statMaxSize);

   IF #NumEvents > #statMaxSize THEN
       #tempScroll_Index_Max := #statMaxSize;
   ELSE
       #tempScroll_Index_Max := #NumEvents;
   END_IF;

   // Statement Section 
   IF #Trigger AND NOT #statTriggerOS THEN
       #statScrollIndex := #statScrollIndex + 1;  // increment the index

       IF  #statScrollIndex > #tempScroll_Index_Max - 1 THEN
               #statScrollIndex := 0;
           END_IF;

      #Msg_Scroll := #In_Events[#statScrollIndex].Message;      // move the message from the UDT_Event structure to string output.  

       #statTriggerOS := TRUE;              // Set the trigger OS bit
   END_IF;

   IF NOT #Trigger AND #statTriggerOS THEN
       #statTriggerOS := FALSE;
   END_IF;

   //  -------------- END OF LOGIC -------------------------
   ENO := TRUE;   // Set the ENO output
END_FUNCTION_BLOCK

FUNCTION_BLOCK "CPG_OEE"   // FB31609, SCL
TITLE = CPG_OEE
{ S7_Optimized_Access := 'TRUE' }
AUTHOR : tech.team.motioncontrol@siemens.com
FAMILY : CPG
VERSION : 1.0
// Support: tech.team.motioncontrol@siemens.com
   VAR_INPUT
      totalProdProcessed : DInt;   // Total Number OF Products Processed
      totalDefectiveProd : DInt;   // Total Number OF Defective Products
      timeSinceLastReset : DInt;   // Total Acumulative TIME since Last RESET
      machineDesignSpeed : Real;   // Machine Design Speed
   END_VAR
   VAR_OUTPUT
      OEERealTimeValue : Real;   // REAL TIME OEE value (availabilty x performance x quality)
      OEEAvailability : Real;   // OEE - Availability value
      OEEPerformance : Real;   // OEE - Performance value
      OEEQuality : Real;   // OEE - Quality value
   END_VAR
   VAR_IN_OUT
      modeCumulativeTimes : Array[0.."LPMLV30_MODES_UPPER_LIM"] of DInt;   // Mode Cummulative Times
   END_VAR
   VAR
      statTotalProdProcessed_In : DInt;   // Initial "TotalProdProcessed" value after accum TIME reset
      statTotalDefectiveProd_In : DInt;   // Initial "TotalDefectiveProcessed" value after accum TIME reset
      statAcumTimeEqualZero : Bool;   // The "TimeSinceLastReset" is = 0 seconds
      statAcumTimeEqualZeroOS : Bool;   // OneShot for "TimeSinceLastReset" is = 0 seconds
   END_VAR
   VAR_TEMP
      tempTimeSinceLastReset : Real;   // used to eliminate divide by zero errors
      tempTotalProducts : Real;   // used to eliminate divide by zero errors
      tempDefectiveProducts : Real;   // used to eliminate divide by zero errors
   END_VAR
BEGIN
   //============================================================================================================
   // SIEMENS AG
   // (c)Copyright 2018 All Rights Reserved
   //------------------------------------------------------------------------------------------------------------
   // Project: CPG Template
   // Tested with: S7-1500 with FW version V2.1
   // Engineering: TIA Portal V14
   // Restrictions: ---
   // Requirements: S7-1500
   // Functionality:  calculate real-time OEE values
   // Support: tech.team.motioncontrol@siemens.com
   //------------------------------------------------------------------------------------------------------------
   // Change log table:
   // Version       Date               Expert in charge    Changes applied
   //  01.00.00     28.02.1012         MP                  Original - using OEE Realtime calculation
   //  01.01.00     04.09.2014         MP                  Added seperate Availabity, Performace, Quality calculation
   //  01.02.00     07.07.2014         MP                  Updated interface FOR new Mode/State FB          
   //  01.02.01     01.02.2016         MP                  Added logic to prevent floating point / divide by zero errors
   //  02.00.00     01.01.2018         MP                  Prepared for CPG Release
   //  02.01.00     29.05.2018         JP                  Adopted to styleguide
   //============================================================================================================
   // Function Block : CPG_OEE
   //============================================================================================================

   // ===========================================================================
   //  Begin the LOGIC section:
   //  
   (* ISA TR88.00.02 Document - 9.1 OEE Definition:
   Overall Equipment Effectiveness (OEE) is a measure comparing how well manufacturing equipment is running compared to the ideal plant. The resulting measurement is expressed as the ratio of the actual
   output of the equipment divided by the maximum possible output of the equipment under ideal conditions. OEE is calculated by multiplying three independently measured values: Availability,
   Performance Rate, and Quality Rate. The fundamental OEE definition is defined as an availability ratio multiplied by a performance ratio multiplied by a quality ratio.

   OEE = Availability x Performance x Quality

   Where each component is defined as the following:
   Availability = Operating Time / Planned Production Time
   Performance = Total Pieces / (Operating Time* Ideal Run Rate)
   Quality = Good Pieces / Total Pieces

   OEE is often displayed as a waterfall object in which the major components of Availability, Performance, and Quality are displayed graphically.
   *)

   // Determine is TimeSinceLastReset value is equal to zero.
   IF  #timeSinceLastReset   = 0 THEN
       #statAcumTimeEqualZero   := TRUE;  // SET the AcumTimeEqualZero bool tag
   ELSE
       #statAcumTimeEqualZero   := FALSE; // RESET the AcumTimeEqualZero bool tag
       #statAcumTimeEqualZeroOS := FALSE; // RESET the AcumTimeEqualZero one-shot bool tag
   END_IF;

   // Update the AcumTimeEqualZeroOS One-Shot bool
   IF #statAcumTimeEqualZero AND NOT #statAcumTimeEqualZeroOS THEN
      #statAcumTimeEqualZeroOS := TRUE;  // Set the One-Shot bool tag
   END_IF;

   // Update the initial product count values after the accum timer value has been reset
   IF #statAcumTimeEqualZeroOS THEN
      #statTotalProdProcessed_In := #totalProdProcessed;
      #statTotalDefectiveProd_In := #totalDefectiveProd;
   END_IF;  

   // Update the TimeSinceLastReset temp. value.  If = 0 (zero) then change to 0.0001 to ensure no divide by zero errors
   IF #timeSinceLastReset = 0 THEN
       #tempTimeSinceLastReset := 0.0001;
   ELSE
       #tempTimeSinceLastReset := DINT_TO_REAL(#timeSinceLastReset);
   END_IF;



   (*  9.1.1 Availability Definition
   Availability is defined as operating time divided by planned production time. The basic concept behind availability is to show the time the machine has been running divided by the time that the
   machine has been planned to run. Typical losses in this area are losses to unplanned maintenance, cleaning, changeovers, and breakdowns.
   * Availability = Operating Time / Planned Production Time Operating Time is defined as the amount of time the machine has been attempting to produce parts.  
   * Planned Production Time is defined as the total amount of time the machine has been scheduled to run. 
   *)
   // Availablity = operating time (attempt to run production) / planned production time
   #OEEAvailability :=   DINT_TO_REAL (#modeCumulativeTimes[1]) / #tempTimeSinceLastReset;
   IF #OEEAvailability > 1.0 THEN #OEEAvailability := 1.0; END_IF;
   IF #OEEAvailability < 0.0 THEN #OEEAvailability := 0.0; END_IF;

   (* 9.1.2 Performance Definition
   Performance is defined as the total number of pieces on which the machine operated divided by the ideal production if a machine ran perfectly for the allocated amount of operating time.
   * Performance = Total Pieces / (Operating Time* Ideal Run Rate).  
   * Total Pieces is defined as good pieces and bad pieces during the production run. This should be linked to the main consumed count of the machine. If a filler, this should be bottles into the filler.
   * Operating Time is defined as the amount of time the machine has been attempting to produce parts. (Same as above)
   * Ideal Run Rate is defined as the ideal rate that the machine can run for the product that is being run on the machine and the way the machine is configured.
   *)
   // Performance = Total Pieces / (Operating Time * Ideal Run Rate / 60)
   #OEEPerformance := (DINT_TO_REAL(#totalProdProcessed - #statTotalProdProcessed_In)) / ((#tempTimeSinceLastReset * #machineDesignSpeed / 60.0));
   IF #OEEPerformance > 1.0 THEN #OEEPerformance := 1.0; END_IF;
   IF #OEEPerformance < 0.0 THEN #OEEPerformance := 0.0; END_IF;

   (*  9.1.3 Quality Definition
   Quality is defined as the total number of good pieces divided by the total number of pieces on which the machine operated.
   * Quality = Good Pieces / Total Pieces
   * Good Pieces is defined as only good pieces processed during the production run. So this is the main production processed count of the machine. If a filler, this should be bottles out of the filler.
   * Total Pieces includes good pieces and bad pieces during the production run. This should be linked to the main consumed count of the machine. 
      If a filler, this should be bottles into the filler. This should be the same count as used in the performance definition.
   *)
   // Quality = Good Piece / Total Piece
   #tempTotalProducts     :=  DINT_TO_REAL(#totalProdProcessed-#statTotalProdProcessed_In);
   #tempDefectiveProducts :=  DINT_TO_REAL(#totalDefectiveProd-#statTotalDefectiveProd_In);

   // Prevent divide by zero errors by checking if Total Products <> 0.0
   IF (#totalProdProcessed - #statTotalProdProcessed_In) = 0 THEN 
       #tempTotalProducts := 0.0001;
   END_IF;

   // Make sure that defective products < total products
   IF #tempDefectiveProducts > #tempTotalProducts THEN
       #tempDefectiveProducts := 0.0;
   END_IF;

   #OEEQuality            := (#tempTotalProducts - #tempDefectiveProducts) / #tempTotalProducts;

   IF #OEEQuality  > 1.0 THEN #OEEQuality  := 1.0; END_IF;
   IF #OEEQuality  < 0.0 THEN #OEEQuality  := 0.0; END_IF;
   IF #tempTotalProducts = 0 THEN
       #OEEQuality := 0.0;
   END_IF;


   #OEERealTimeValue := #OEEAvailability * #OEEPerformance * #OEEQuality;

   //  -------------- END OF LOGIC -------------------------
   ENO := TRUE;   // Set the ENO output
END_FUNCTION_BLOCK

